text list "Banner_WarnMsg2": 0 '**Local Message Display**'; 1 '~Safety Task Unlocked WB2[0].1'; 2 '~Safety Signature Mismatch WB2[0].2'; 3 '~PLC Battery Bad Or Missing WB2[0].3'; 4 '~Lube System Faulted WB2[0].4'; 5 '~Lube System Cycling WB2[0].5'; 6 '~Lube Level Low WB2[0].6'; 7 '~Spare WB2[0].7'; 8 '~Spare WB2[0].8'; 9 '~Spare WB2[0].9'; 10 '~Main Air Filter Dirty WB2[0].10'; 11 '~Main Water Filter Not OK WB2[0].11'; 12 '~Spare WB2[0].12'; 13 '~Spare WB2[0].13'; 14 '~Spare WB2[0].14'; 15 '~Spare WB2[0].15'; 16 '~Spare WB2[0].16'; 17 '~Spare WB2[0].17'; 18 '~Spare WB2[0].18'; 19 '~Spare WB2[0].19'; 20 '~Spare WB2[0].20'; 21 '~Spare WB2[0].21'; 22 '~Spare WB2[0].22'; 23 '~Spare WB2[0].23'; 24 '~Spare WB2[0].24'; 25 '~Spare WB2[0].25'; 26 '~Spare WB2[0].26'; 27 '~Spare WB2[0].27'; 28 '~Spare WB2[0].28'; 29 '~Spare WB2[0].29'; 30 '~Spare WB2[0].30'; 31 '~Spare WB2[0].31'; 32 '~Sxxx-xxx - Prev Station Exit Lt Scrn Fault - See Prev Station PV WB2[1].0'; 33 '~Sxxx-xxx - Next Station Exit Lt Scrn Fault - See Next Station PV WB2[1].1'; 34 '~Sxxx-xxx - Prev Station Robot In Teach - See Prev Station PV WB2[1].2'; 35 '~Sxxx-xxx - Next Station Robot In Teach - See Next Station PV WB2[1].3'; 36 '~Spare WB2[1].4'; 37 '~Spare WB2[1].5'; 38 '~Sxxx-xxx - Facilities Gate Logic Not Rst - See Facilities Ctrl Pnl WB2[1].6'; 39 '~Spare WB2[1].7'; 40 '~Spare WB2[1].8'; 41 '~Sxxx-xxx - Other Control Zone Fault Present WB2[1].9'; 42 '~Spare WB2[1].10'; 43 '~Spare WB2[1].11'; 44 '~Safety Instruction Warning - Go To Safety Instruction Screen WB2[1].12'; 45 '~Safety Instruction Fault Active - Go To Safety Instuction Screen WB2[1].13'; 46 '~Spare WB2[1].14'; 47 '~Spare WB2[1].15'; 48 '~Spare WB2[1].16'; 49 '~Spare WB2[1].17'; 50 '~Spare WB2[1].18'; 51 '~Spare WB2[1].19'; 52 '~Spare WB2[1].20'; 53 '~Sxxx-xxx Consumed Safety I/O Intlks Not Running-See Source PLC WB2[1].21'; 54 '~Sxxx-xxx Consumed Standard I/O Intlks Not Running-See Source PLC WB2[1].22'; 55 '~Sxxx-xxx Consumed Safety I/O Intlks Not Running-See Source PLC WB2[1].23'; 56 '~Sxxx-xxx Consumed Standard I/O Intlks Not Running-See Source PLC WB2[1].24'; 57 '~Sxxx-xxx Consumed Safety I/O Intlks Not Running-See Source PLC WB2[1].25'; 58 '~Sxxx-xxx Consumed Standard I/O Intlks Not Running-See Source PLC WB2[1].26'; 59 '~Sxxx-xxx Consumed Safety I/O Intlks Not Running-See Source PLC WB2[1].27'; 60 '~Sxxx-xxx Consumed Standard I/O Intlks Not Running-See Source PLC WB2[1].28'; 61 '~Spare WB2[1].29'; 62 '~Spare WB2[1].30'; 63 '~Spare WB2[1].31'; 64 '~Sxxx - xxx E-Stop Depressed - See Station Panel WB2[2].0'; 65 '~Sxxx - xxx E-Stop Circuit Not Reset - Depress Enable Outputs PB WB2[2].1'; 66 '~Sxxx - xxx Safety Gate Open - See Station Panel WB2[2].2'; 67 '~Sxxx - xxx Safety Gate Circuit Not Reset - Depress Gate Reset PB WB2[2].3'; 68 '~Sxxx - xxx Access Or Entry/Exit Light Screen Fault - See Stn Panel WB2[2].4'; 69 '~Sxxx - xxx Robot In Teach - See Station Panel WB2[2].5'; 70 '~Sxxx - xxx Not Ready For Auto - See Station Panel WB2[2].6'; 71 '~Sxxx - xxx Auto Repeat Not Selected - See Station Panel WB2[2].7'; 72 '~Sxxx - xxx Faulted - See Station Panel WB2[2].8'; 73 '~Spare WB2[2].9'; 74 '~Spare WB2[2].10'; 75 '~Spare WB2[2].11'; 76 '~Spare WB2[2].12'; 77 '~Spare WB2[2].13'; 78 '~Spare WB2[2].14'; 79 '~Spare WB2[2].15'; 80 '~Sxxx - xxx E-Stop Depressed - See Station Panel WB2[2].16'; 81 '~Sxxx - xxx E-Stop Circuit Not Reset - Depress Enable Outputs PB WB2[2].17'; 82 '~Sxxx - xxx Safety Gate Open - See Station Panel WB2[2].18'; 83 '~Sxxx - xxx Safety Gate Circuit Not Reset - Depress Gate Reset PB WB2[2].19'; 84 '~Sxxx - xxx Access Or Entry/Exit Light Screen Fault - See Stn Panel WB2[2].20'; 85 '~Sxxx - xxx Robot In Teach - See Station Panel WB2[2].21'; 86 '~Sxxx - xxx Not Ready For Auto - See Station Panel WB2[2].22'; 87 '~Sxxx - xxx Auto Repeat Not Selected - See Station Panel WB2[2].23'; 88 '~Sxxx - xxx Faulted - See Station Panel WB2[2].24'; 89 '~Spare WB2[2].25'; 90 '~Spare WB2[2].26'; 91 '~Spare WB2[2].27'; 92 '~Spare WB2[2].28'; 93 '~Spare WB2[2].29'; 94 '~Spare WB2[2].30'; 95 '~Spare WB2[2].31'; 96 '~Sxxx - xxx E-Stop Depressed - See Station Panel WB2[3].0'; 97 '~Sxxx - xxx E-Stop Circuit Not Reset - Depress Enable Outputs PB WB2[3].1'; 98 '~Sxxx - xxx Safety Gate Open - See Station Panel WB2[3].2'; 99 '~Sxxx - xxx Safety Gate Circuit Not Reset - Depress Gate Reset PB WB2[3].3'; 100 '~Sxxx - xxx Access Or Entry/Exit Light Screen Fault - See Stn Panel WB2[3].4'; 101 '~Sxxx - xxx Robot In Teach - See Station Panel WB2[3].5'; 102 '~Sxxx - xxx Not Ready For Auto - See Station Panel WB2[3].6'; 103 '~Sxxx - xxx Auto Repeat Not Selected - See Station Panel WB2[3].7'; 104 '~Sxxx - xxx Faulted - See Station Panel WB2[3].8'; 105 '~Spare WB2[3].9'; 106 '~Spare WB2[3].10'; 107 '~Spare WB2[3].11'; 108 '~Spare WB2[3].12'; 109 '~Spare WB2[3].13'; 110 '~Spare WB2[3].14'; 111 '~Spare WB2[3].15'; 112 '~Sxxx - xxx E-Stop Depressed - See Station Panel WB2[3].16'; 113 '~Sxxx - xxx E-Stop Circuit Not Reset - Depress Enable Outputs PB WB2[3].17'; 114 '~Sxxx - xxx Safety Gate Open - See Station Panel WB2[3].18'; 115 '~Sxxx - xxx Safety Gate Circuit Not Reset - Depress Gate Reset PB WB2[3].19'; 116 '~Sxxx - xxx Access Or Entry/Exit Light Screen Fault - See Stn Panel WB2[3].20'; 117 '~Sxxx - xxx Robot In Teach - See Station Panel WB2[3].21'; 118 '~Sxxx - xxx Not Ready For Auto - See Station Panel WB2[3].22'; 119 '~Sxxx - xxx Auto Repeat Not Selected - See Station Panel WB2[3].23'; 120 '~Sxxx - xxx Faulted - See Station Panel WB2[3].24'; 121 '~Spare WB2[3].25'; 122 '~Spare WB2[3].26'; 123 '~Spare WB2[3].27'; 124 '~Spare WB2[3].28'; 125 '~Spare WB2[3].29'; 126 '~Spare WB2[3].30'; 127 '~Spare WB2[3].31'; 128 '~Sxxx - xxx E-Stop Depressed - See Station Panel WB2[4].0'; 129 '~Sxxx - xxx E-Stop Circuit Not Reset - Depress Enable Outputs PB WB2[4].1'; 130 '~Sxxx - xxx Safety Gate Open - See Station Panel WB2[4].2'; 131 '~Sxxx - xxx Safety Gate Circuit Not Reset - Depress Gate Reset PB WB2[4].3'; 132 '~Sxxx - xxx Access Or Entry/Exit Light Screen Fault WB2[4].4'; 133 '~Sxxx - xxx Robot In Teach - See Station Panel WB2[4].5'; 134 '~Sxxx - xxx Not Ready For Auto - See Station Panel WB2[4].6'; 135 '~Sxxx - xxx Auto Repeat Not Selected - See Station Panel WB2[4].7'; 136 '~Sxxx - xxx Faulted - See Station Panel WB2[4].8'; 137 '~Spare WB2[4].9'; 138 '~Spare WB2[4].10'; 139 '~Spare WB2[4].11'; 140 '~Spare WB2[4].12'; 141 '~Spare WB2[4].13'; 142 '~Spare WB2[4].14'; 143 '~Spare WB2[4].15'; 144 '~Spare WB2[4].16'; 145 '~Spare WB2[4].17'; 146 '~Spare WB2[4].18'; 147 '~Spare WB2[4].19'; 148 '~Spare WB2[4].20'; 149 '~Spare WB2[4].21'; 150 '~Spare WB2[4].22'; 151 '~Spare WB2[4].23'; 152 '~Spare WB2[4].24'; 153 '~Spare WB2[4].25'; 154 '~Spare WB2[4].26'; 155 '~Spare WB2[4].27'; 156 '~Spare WB2[4].28'; 157 '~Spare WB2[4].29'; 158 '~Spare WB2[4].30'; 159 '~Spare WB2[4].31'; 160 '~S002 Safety Gate Logic Not Reset - Depress Gate Reset PB WB2[5].0'; 161 '~Spare WB2[5].1'; 162 '~Spare WB2[5].2'; 163 '~Spare WB2[5].3'; 164 '~S002 Ready For Automatic Depress Auto PB WB2[5].4'; 165 '~S002 Master Logic Not Reset Depress Enable Ouputs PB WB2[5].5'; 166 '~S002 Not Ready For Automatic WB2[5].6'; 167 '~S002 Auto Repeat Not Selected - See Utility Screen WB2[5].7'; 168 '~Spare WB2[5].8'; 169 '~Spare WB2[5].9'; 170 '~S002 Service Side Light Screen Not Reset - Depress Cycle Start PB WB2[5].10'; 171 '~S002 Remote Side Light Screen Not Reset - Depress Cycle Start PB WB2[5].11'; 172 '~Spare WB2[5].12'; 173 '~Spare WB2[5].13'; 174 '~Spare WB2[5].14'; 175 '~Spare WB2[5].15'; 176 '~Spare WB2[5].16'; 177 '~Spare WB2[5].17'; 178 '~Spare WB2[5].18'; 179 '~Spare WB2[5].19'; 180 '~Spare WB2[5].20'; 181 '~Spare WB2[5].21'; 182 '~Spare WB2[5].22'; 183 '~Spare WB2[5].23'; 184 '~S002 Service Side Model 1 Prycheck Selected WB2[5].24'; 185 '~S002 Remote Side Model 1 Prycheck Selected WB2[5].25'; 186 '~S002 Service Side Model 2 Prycheck Selected WB2[5].26'; 187 '~S002 Remote Side Model 2 Prycheck Selected WB2[5].27'; 188 '~Spare WB2[5].28'; 189 '~Spare WB2[5].29'; 190 '~Spare WB2[5].30'; 191 '~Spare WB2[5].31'; 192 '~Spare WB2[6].0'; 193 '~Spare WB2[6].1'; 194 '~S002 Oper #1 Light Screen Not Reset - Press Cycle Start PB WB2[6].2'; 195 '~S002 Oper #2 Light Screen Not Reset - Press Cycle Start PB WB2[6].3'; 196 '~S002CV# Oper #1 Lt Screen Not Reset - Press Cycle Start PB WB2[6].4'; 197 '~S002CV# Oper #2 Lt Screen Not Reset - Press Cycle Start PB WB2[6].5'; 198 '~Spare WB2[6].6'; 199 '~Spare WB2[6].7'; 200 '~Spare WB2[6].8'; 201 '~Spare WB2[6].9'; 202 '~S002 Operator #1 Cycle Over Time WB2[6].10'; 203 '~S002 Operator #2 Cycle Overtime WB2[6].11'; 204 '~S002TT1 Operator #1 Cycle Over Time WB2[6].12'; 205 '~S003TL1 Operator #1 Cycle Over Time WB2[6].13'; 206 '~Spare WB2[6].14'; 207 '~Spare WB2[6].15'; 208 '~Spare WB2[6].16'; 209 '~Spare WB2[6].17'; 210 '~Spare WB2[6].18'; 211 '~Spare WB2[6].19'; 212 '~Spare WB2[6].20'; 213 '~Spare WB2[6].21'; 214 '~Spare WB2[6].22'; 215 '~Spare WB2[6].23'; 216 '~Spare WB2[6].24'; 217 '~Spare WB2[6].25'; 218 '~Spare WB2[6].26'; 219 '~Spare WB2[6].27'; 220 '~Spare WB2[6].28'; 221 '~Spare WB2[6].29'; 222 '~Spare WB2[6].30'; 223 '~Spare WB2[6].31'; 224 '~PDPES1 - PDP EtherNet Switch Port At Half Duplex WB2[7].0'; 225 '~PDPES1 - PDP EtherNet Switch Configuration Changes Not Saved WB2[7].1'; 226 '~PDPES1 - PDP EtherNet Switch Configuration Changed WB2[7].2'; 227 '~PDPES1 - PDP EtherNet Switch Port With Excessive Errors WB2[7].3'; 228 '~PDPES1 - PDP EtherNet Switch Port With Utilization Warning WB2[7].4'; 229 '~PDPES1 - PDP EtherNet Switch Changes Require Reboot WB2[7].5'; 230 '~Spare WB2[7].6'; 231 '~Spare WB2[7].7'; 232 '~MPES1 - Main Panel EtherNet Switch Port At Half Duplex WB2[7].8'; 233 '~MPES1 - Main Panel EtherNet Switch Configuration Changes Not Saved WB2[7].9'; 234 '~MPES1 - Main Panel EtherNet Switch Configuration Changed WB2[7].10'; 235 '~MPES1 - Main Panel EtherNet Switch Port With Excessive Errors WB2[7].11'; 236 '~MPES1 - Main Panel EtherNet Switch Port With Utilization Warning WB2[7].12'; 237 '~MPES1 - Main Panel EtherNet Switch Changes Require Reboot WB2[7].13'; 238 '~Spare WB2[7].14'; 239 '~Spare WB2[7].15'; 240 '~MPES2 - Main Panel EtherNet Switch Port At Half Duplex WB2[7].16'; 241 '~MPES2 - Main Panel EtherNet Switch Configuration Changes Not Saved WB2[7].17'; 242 '~MPES2 - Main Panel EtherNet Switch Configuration Changed WB2[7].18'; 243 '~MPES2 - Main Panel EtherNet Switch Port With Excessive Errors WB2[7].19'; 244 '~MPES2 - Main Panel EtherNet Switch Port With Utilization Warning WB2[7].20'; 245 '~MPES2 - Main Panel EtherNet Switch Changes Require Reboot WB2[7].21'; 246 '~Spare WB2[7].22'; 247 '~Spare WB2[7].23'; 248 '~MPES3 - Main Panel EtherNet Switch Port At Half Duplex WB2[7].24'; 249 '~MPES3 - Main Panel EtherNet Switch Configuration Changes Not Saved WB2[7].25'; 250 '~MPES3 - Main Panel EtherNet Switch Configuration Changed WB2[7].26'; 251 '~MPES3 - Main Panel EtherNet Switch Port With Excessive Errors WB2[7].27'; 252 '~MPES3 - Main Panel EtherNet Switch Port With Utilization Warning WB2[7].28'; 253 '~MPES3 - Main Panel EtherNet Switch Changes Require Reboot WB2[7].29'; 254 '~Spare WB2[7].30'; 255 '~Spare WB2[7].31'; 256 '~PV3ES1 - PV3 EtherNet Switch Port At Half Duplex WB2[8].0'; 257 '~PV3ES1 - PV3 EtherNet Switch Configuration Changes Not Saved WB2[8].1'; 258 '~PV3ES1 - PV3 EtherNet Switch Configuration Changed WB2[8].2'; 259 '~PV3ES1 - PV3 EtherNet Switch Port With Excessive Errors WB2[8].3'; 260 '~PV3ES1 - PV3 EtherNet Switch Port With Utilization Warning WB2[8].4'; 261 '~PV3ES1 - PV3 EtherNet Switch Changes Require Reboot WB2[8].5'; 262 '~Spare WB2[8].6'; 263 '~Spare WB2[8].7'; 264 '~PV4ES1 - PV4 EtherNet Switch Port At Half Duplex WB2[8].8'; 265 '~PV4ES1 - PV4 EtherNet Switch Configuration Changes Not Saved WB2[8].9'; 266 '~PV4ES1 - PV4 EtherNet Switch Configuration Changed WB2[8].10'; 267 '~PV4ES1 - PV4 EtherNet Switch Port With Excessive Errors WB2[8].11'; 268 '~PV4ES1 - PV4 EtherNet Switch Port With Utilization Warning WB2[8].12'; 269 '~PV4ES1 - PV4 EtherNet Switch Changes Require Reboot WB2[8].13'; 270 '~Spare WB2[8].14'; 271 '~Spare WB2[8].15'; 272 '~ES3ES1 - ES3 EtherNet Switch Port At Half Duplex WB2[8].16'; 273 '~ES3ES1 - ES3 EtherNet Switch Configuration Changes Not Saved WB2[8].17'; 274 '~ES3ES1 - ES3 EtherNet Switch Configuration Changed WB2[8].18'; 275 '~ES3ES1 - ES3 EtherNet Switch Port With Excessive Errors WB2[8].19'; 276 '~ES3ES1 - ES3 EtherNet Switch Port With Utilization Warning WB2[8].20'; 277 '~ES3ES1 - ES3 EtherNet Switch Changes Require Reboot WB2[8].21'; 278 '~Spare WB2[8].22'; 279 '~Spare WB2[8].23'; 280 '~ES4ES1 - ES4 EtherNet Switch Port At Half Duplex WB2[8].24'; 281 '~ES4ES1 - ES4 EtherNet Switch Configuration Changes Not Saved WB2[8].25'; 282 '~ES4ES1 - ES4 EtherNet Switch Configuration Changed WB2[8].26'; 283 '~ES4ES1 - ES4 EtherNet Switch Port With Excessive Errors WB2[8].27'; 284 '~ES4ES1 - ES4 EtherNet Switch Port With Utilization Warning WB2[8].28'; 285 '~ES4ES1 - ES4 EtherNet Switch Changes Require Reboot WB2[8].29'; 286 '~Spare WB2[8].30'; 287 '~Spare WB2[8].31'; 288 '~Spare WB2[9].0'; 289 '~Spare WB2[9].1'; 290 '~Spare WB2[9].2'; 291 '~Spare WB2[9].3'; 292 '~Spare WB2[9].4'; 293 '~Spare WB2[9].5'; 294 '~Spare WB2[9].6'; 295 '~Spare WB2[9].7'; 296 '~Spare WB2[9].8'; 297 '~Spare WB2[9].9'; 298 '~Spare WB2[9].10'; 299 '~Spare WB2[9].11'; 300 '~Spare WB2[9].12'; 301 '~Spare WB2[9].13'; 302 '~Spare WB2[9].14'; 303 '~Spare WB2[9].15'; 304 '~Spare WB2[9].16'; 305 '~Spare WB2[9].17'; 306 '~Spare WB2[9].18'; 307 '~Spare WB2[9].19'; 308 '~Spare WB2[9].20'; 309 '~Spare WB2[9].21'; 310 '~Spare WB2[9].22'; 311 '~Spare WB2[9].23'; 312 '~Spare WB2[9].24'; 313 '~Spare WB2[9].25'; 314 '~Spare WB2[9].26'; 315 '~Spare WB2[9].27'; 316 '~Spare WB2[9].28'; 317 '~Spare WB2[9].29'; 318 '~Spare WB2[9].30'; 319 '~Spare WB2[9].31'; 320 '~S001R09 Waiting Zone #1 Not Clear WB2[10].0'; 321 '~S001R09 Waiting Zone #2 Not Clear WB2[10].1'; 322 '~S001R09 Waiting Zone #3 Not Clear WB2[10].2'; 323 '~S001R09 Waiting Zone #4 Not Clear WB2[10].3'; 324 '~S001R09 Waiting Zone #5 Not Clear WB2[10].4'; 325 '~S001R09 Waiting Zone #6 Not Clear WB2[10].5'; 326 '~S001R09 Waiting Zone #7 Not Clear WB2[10].6'; 327 '~S001R09 Waiting Zone #8 Not Clear WB2[10].7'; 328 '~S001R09 Waiting Zone #9 Not Clear WB2[10].8'; 329 '~S001R09 Waiting Zone #10 Not Clear WB2[10].9'; 330 '~S001R09 Waiting Zone #11 Not Clear WB2[10].10'; 331 '~S001R09 Waiting Zone #12 Not Clear WB2[10].11'; 332 '~S001R09 Waiting Zone #13 Not Clear WB2[10].12'; 333 '~S001R09 Waiting Zone #14 Not Clear WB2[10].13'; 334 '~S001R09 Waiting Tip Dress Zone #1 Not Clear WB2[10].14'; 335 '~S001R09 Waiting Tip Dress Zone #2 Not Clear WB2[10].15'; 336 '~S001R09 Adjacent Robot xx-xx In Teach WB2[10].16'; 337 '~S001R09 Adjacent Robot xx-xx In Teach WB2[10].17'; 338 '~S001R09 Adjacent Robot xx-xx In Teach WB2[10].18'; 339 '~S001R09 Adjacent Robot xx-xx In Teach WB2[10].19'; 340 '~S001R09 Adjacent Robot xx-xx In Teach WB2[10].20'; 341 '~S001R09 Adjacent Robot xx-xx In Teach WB2[10].21'; 342 '~S001R09 Adjacent Robot xx-xx In Teach WB2[10].22'; 343 '~S001R09 Adjacent Robot xx-xx In Teach WB2[10].23'; 344 '~S001R09 Adjacent Robot xx-xx In Teach WB2[10].24'; 345 '~S001R09 Adjacent Robot xx-xx In Teach WB2[10].25'; 346 '~Spare WB2[10].26'; 347 '~Spare WB2[10].27'; 348 '~Spare WB2[10].28'; 349 '~S001R09 Robot Not Clear Of Fixture WB2[10].29'; 350 '~Spare WB2[10].30'; 351 '~Spare WB2[10].31'; 352 '~Spare WB2[11].0'; 353 '~Spare WB2[11].1'; 354 '~Spare WB2[11].2'; 355 '~Spare WB2[11].3'; 356 '~Spare WB2[11].4'; 357 '~Spare WB2[11].5'; 358 '~Spare WB2[11].6'; 359 '~Spare WB2[11].7'; 360 '~Spare WB2[11].8'; 361 '~Spare WB2[11].9'; 362 '~Spare WB2[11].10'; 363 '~Spare WB2[11].11'; 364 '~Spare WB2[11].12'; 365 '~Spare WB2[11].13'; 366 '~Spare WB2[11].14'; 367 '~Spare WB2[11].15'; 368 '~Spare WB2[11].16'; 369 '~Spare WB2[11].17'; 370 '~Spare WB2[11].18'; 371 '~Spare WB2[11].19'; 372 '~Spare WB2[11].20'; 373 '~Spare WB2[11].21'; 374 '~Spare WB2[11].22'; 375 '~Spare WB2[11].23'; 376 '~Spare WB2[11].24'; 377 '~Spare WB2[11].25'; 378 '~Spare WB2[11].26'; 379 '~Spare WB2[11].27'; 380 '~Spare WB2[11].28'; 381 '~Spare WB2[11].29'; 382 '~Spare WB2[11].30'; 383 '~Spare WB2[11].31'; 384 '~S001R09 Cycle Overtime WB2[12].0'; 385 '~S001R09 In Bypass WB2[12].1'; 386 '~S001R09 Battery Low WB2[12].2'; 387 '~S001R09 Servo Over Torque WB2[12].3'; 388 '~S001R09 Process Retry In Progress WB2[12].4'; 389 '~Spare WB2[12].5'; 390 '~S001R09 Robot Edit Occurred Ext App WB2[12].6'; 391 '~S001R09 Robot Input Simmed WB2[12].7'; 392 '~S001R09 Robot Output Simmed WB2[12].8'; 393 '~Spare WB2[12].9'; 394 '~Spare WB2[12].10'; 395 '~Spare WB2[12].11'; 396 '~Spare WB2[12].12'; 397 '~Spare WB2[12].13'; 398 '~Spare WB2[12].14'; 399 '~Spare WB2[12].15'; 400 '~S001R09F1B1.M.ModuleFlt - Externa App 1 I/O Module Warning WB2[12].16'; 401 '~S001R09F2B1.M.ModuleFlt - Externa App 2 I/O Module Warning WB2[12].17'; 402 '~S001R09F3B1.M.ModuleFlt - Externa App 3 I/O Module Warning WB2[12].18'; 403 '~Spare WB2[12].19'; 404 '~Spare WB2[12].20'; 405 '~Spare WB2[12].21'; 406 '~Spare WB2[12].22'; 407 '~Spare WB2[12].23'; 408 '~S001R09ES1 - S001R09 EtherNet Switch Port At Half Duplex WB2[12].24'; 409 '~S001R09ES1 - S001R09 EtherNet Switch Config Changes Not Saved WB2[12].25'; 410 '~S001R09ES1 - S001R09 EtherNet Switch Configuration Changed WB2[12].26'; 411 '~S001R09ES1 - S001R09 EtherNet Switch Port With Excessive Errors WB2[12].27'; 412 '~S001R09ES1 - S001R09 EtherNet Switch Port With Utilization Warning WB2[12].28'; 413 '~S001R09ES1 - S001R09 EtherNet Switch Changes Require Reboot WB2[12].29'; 414 '~Spare WB2[12].30'; 415 '~Spare WB2[12].31'; 416 '~Spare WB2[13].0'; 417 '~Spare WB2[13].1'; 418 '~S001R09 Servo Gun Tip Calib Request 1 WB2[13].2'; 419 '~S001R09 I-Available Warning 1 WB2[13].3'; 420 '~S001R09 Tip Dress Motor 1 Fault Bypassed WB2[13].4'; 421 '~S001R09 Tip Change Notice 1 WB2[13].5'; 422 '~S001R09 Bypass Tip Dresser 1 Selected WB2[13].6'; 423 '~S001R09 Auto Tip Changer Low 1 WB2[13].7'; 424 '~S001R09 Auto Tip Changer Empty 1 WB2[13].8'; 425 '~S001R09 Tip Wear Ratio Warning 1 - Touch Up Tip Dress Program WB2[13].9'; 426 '~S001R09 Stud Weld 1 Maintenance Reqd WB2[13].10'; 427 '~S001R09 Stud Weld 1 Low Stud Warning WB2[13].11'; 428 '~Spare WB2[13].12'; 429 '~S001R09 Rivet 1 Low Rivet Warning WB2[13].13'; 430 '~S001R09 Rivet 1 - Skip Once Initiated from Robot TP WB2[13].14'; 431 '~S001R09 Rivet 1 - Skip Remaining Initiated from Robot TP WB2[13].15'; 432 '~S001R09 Rivet 1 Preventive Maintenace Required WB2[13].16'; 433 '~S001R09 Rivet 1 Magazine Low WB2[13].17'; 434 '~S001R09 Tip Change 1 Bypassed WB2[13].18'; 435 '~S001R09 Mig Weld Fluid Level Low WB2[13].19'; 436 '~S001R09 Weld Ctrlr 1 Adaptive Mode Is Disabled WB2[13].20'; 437 '~S001R09 Tip Cutter 1 Warning WB2[13].21'; 438 '~S001R09 Rivet 1 Tape-Cut Required WB2[13].22'; 439 '~S001R09 Wire Feeder Motor Over Current WB2[13].23'; 440 '~Spare WB2[13].24'; 441 '~S001R09 Sealer Ctrlr 1 Minor Fault WB2[13].25'; 442 '~S001R09 Sealer Ctrlr 1 Required Rezeroing WB2[13].26'; 443 '~S001R09 Loaded To Average WB2[13].27'; 444 '~S001R09 Vision Process Aborted WB2[13].28'; 445 '~S001R09 Vision System Trending WB2[13].29'; 446 '~S001R09 Vision Out Of Tolerance WB2[13].30'; 447 '~Spare WB2[13].31'; 448 '~Spare WB2[14].0'; 449 '~Spare WB2[14].1'; 450 '~S001R09 Servo Gun Tip Calib Request 2 WB2[14].2'; 451 '~S001R09 I-Available Warning 2 WB2[14].3'; 452 '~S001R09 Tip Dress Motor 2 Fault Bypassed WB2[14].4'; 453 '~S001R09 Tip Change Notice 2 WB2[14].5'; 454 '~S001R09 Bypass Tip Dresser 2 Selected WB2[14].6'; 455 '~S001R09 Auto Tip Changer Low 2 WB2[14].7'; 456 '~S001R09 Auto Tip Changer Empty 2 WB2[14].8'; 457 '~S001R09 Tip Wear Ratio Warning 2 - Touch Up Tip Dress Program WB2[14].9'; 458 '~S001R09 Stud Weld 2 Maintenance Reqd WB2[14].10'; 459 '~S001R09 Stud Weld 2 Low Stud Warning WB2[14].11'; 460 '~Spare WB2[14].12'; 461 '~S001R09 Rivet 2 Low Rivet Warning WB2[14].13'; 462 '~S001R09 Rivet 2 - Skip Once Initiated from Robot TP WB2[14].14'; 463 '~S001R09 Rivet 2 - Skip Remaining Initiated from Robot TP WB2[14].15'; 464 '~S001R09 Rivet 2 Preventive Maintenace Required WB2[14].16'; 465 '~S001R09 Rivet 2 Magazine Low WB2[14].17'; 466 '~S001R09 Tip Change 2 Bypassed WB2[14].18'; 467 '~S001R09 Laser Dirty Glass Warning WB2[14].19'; 468 '~S001R09 Weld Ctrlr 2 Adaptive Mode Is Disabled WB2[14].20'; 469 '~S001R09 Tip Cutter 2 Warning WB2[14].21'; 470 '~S001R09 Rivet 2 Tape-Cut Required WB2[14].22'; 471 '~S001R09 Mig Tip Nozzel Replacement Warning WB2[14].23'; 472 '~S001R09 Mig Tip Nozzel Replacement Required WB2[14].24'; 473 '~S001R09 Sealer Ctrlr 2 Minor Fault WB2[14].25'; 474 '~S001R09 Sealer Ctrlr 2 Required Rezeroing WB2[14].26'; 475 '~S001R09 Mig Barrel Replacement Warning WB2[14].27'; 476 '~S001R09 Mig Barrel Replacement Required WB2[14].28'; 477 '~S001R09 In Touch Up Mode WB2[14].29'; 478 '~S001R09 Touch Up Mode Not Enabled WB2[14].30'; 479 '~Spare WB2[14].31'; 480 '~S001R09 Laser Controller Fault WB2[15].0'; 481 '~S001R09 Laser Dirty Glass Warning WB2[15].1'; 482 '~S001R09 Laser Warning WB2[15].2'; 483 '~Spare WB2[15].3'; 484 '~Spare WB2[15].4'; 485 '~Spare WB2[15].5'; 486 '~Spare WB2[15].6'; 487 '~Spare WB2[15].7'; 488 '~Spare WB2[15].8'; 489 '~Spare WB2[15].9'; 490 '~Spare WB2[15].10'; 491 '~Spare WB2[15].11'; 492 '~Spare WB2[15].12'; 493 '~Spare WB2[15].13'; 494 '~Spare WB2[15].14'; 495 '~Spare WB2[15].15'; 496 '~Spare WB2[15].16'; 497 '~Spare WB2[15].17'; 498 '~Spare WB2[15].18'; 499 '~Spare WB2[15].19'; 500 '~Spare WB2[15].20'; 501 '~Spare WB2[15].21'; 502 '~Spare WB2[15].22'; 503 '~Spare WB2[15].23'; 504 '~Spare WB2[15].24'; 505 '~Spare WB2[15].25'; 506 '~Spare WB2[15].26'; 507 '~Spare WB2[15].27'; 508 '~Spare WB2[15].28'; 509 '~Spare WB2[15].29'; 510 '~Spare WB2[15].30'; 511 '~Spare WB2[15].31'; 512 '~Spare WB2[16].0'; 513 '~Spare WB2[16].1'; 514 '~Spare WB2[16].2'; 515 '~Spare WB2[16].3'; 516 '~Spare WB2[16].4'; 517 '~Spare WB2[16].5'; 518 '~Spare WB2[16].6'; 519 '~Spare WB2[16].7'; 520 '~Spare WB2[16].8'; 521 '~Spare WB2[16].9'; 522 '~Spare WB2[16].10'; 523 '~Spare WB2[16].11'; 524 '~Spare WB2[16].12'; 525 '~Spare WB2[16].13'; 526 '~Spare WB2[16].14'; 527 '~Spare WB2[16].15'; 528 '~Spare WB2[16].16'; 529 '~Spare WB2[16].17'; 530 '~Spare WB2[16].18'; 531 '~Spare WB2[16].19'; 532 '~Spare WB2[16].20'; 533 '~Spare WB2[16].21'; 534 '~Spare WB2[16].22'; 535 '~Spare WB2[16].23'; 536 '~Spare WB2[16].24'; 537 '~Spare WB2[16].25'; 538 '~Spare WB2[16].26'; 539 '~Spare WB2[16].27'; 540 '~Spare WB2[16].28'; 541 '~Spare WB2[16].29'; 542 '~Spare WB2[16].30'; 543 '~Spare WB2[16].31'; 544 '~Spare WB2[17].0'; 545 '~Spare WB2[17].1'; 546 '~Spare WB2[17].2'; 547 '~Spare WB2[17].3'; 548 '~Spare WB2[17].4'; 549 '~Spare WB2[17].5'; 550 '~Spare WB2[17].6'; 551 '~Spare WB2[17].7'; 552 '~Spare WB2[17].8'; 553 '~Spare WB2[17].9'; 554 '~Spare WB2[17].10'; 555 '~Spare WB2[17].11'; 556 '~Spare WB2[17].12'; 557 '~Spare WB2[17].13'; 558 '~Spare WB2[17].14'; 559 '~Spare WB2[17].15'; 560 '~Spare WB2[17].16'; 561 '~Spare WB2[17].17'; 562 '~Spare WB2[17].18'; 563 '~Spare WB2[17].19'; 564 '~Spare WB2[17].20'; 565 '~Spare WB2[17].21'; 566 '~Spare WB2[17].22'; 567 '~Spare WB2[17].23'; 568 '~Spare WB2[17].24'; 569 '~Spare WB2[17].25'; 570 '~Spare WB2[17].26'; 571 '~Spare WB2[17].27'; 572 '~Spare WB2[17].28'; 573 '~Spare WB2[17].29'; 574 '~Spare WB2[17].30'; 575 '~Spare WB2[17].31'; 576 '~S001R10 Waiting Zone #1 Not Clear WB2[18].0'; 577 '~S001R10 Waiting Zone #2 Not Clear WB2[18].1'; 578 '~S001R10 Waiting Zone #3 Not Clear WB2[18].2'; 579 '~S001R10 Waiting Zone #4 Not Clear WB2[18].3'; 580 '~S001R10 Waiting Zone #5 Not Clear WB2[18].4'; 581 '~S001R10 Waiting Zone #6 Not Clear WB2[18].5'; 582 '~S001R10 Waiting Zone #7 Not Clear WB2[18].6'; 583 '~S001R10 Waiting Zone #8 Not Clear WB2[18].7'; 584 '~S001R10 Waiting Zone #9 Not Clear WB2[18].8'; 585 '~S001R10 Waiting Zone #10 Not Clear WB2[18].9'; 586 '~S001R10 Waiting Zone #11 Not Clear WB2[18].10'; 587 '~S001R10 Waiting Zone #12 Not Clear WB2[18].11'; 588 '~S001R10 Waiting Zone #13 Not Clear WB2[18].12'; 589 '~S001R10 Waiting Zone #14 Not Clear WB2[18].13'; 590 '~S001R10 Waiting Tip Dress Zone #1 Not Clear WB2[18].14'; 591 '~S001R10 Waiting Tip Dress Zone #2 Not Clear WB2[18].15'; 592 '~S001R10 Adjacent Robot xx-xx In Teach WB2[18].16'; 593 '~S001R10 Adjacent Robot xx-xx In Teach WB2[18].17'; 594 '~S001R10 Adjacent Robot xx-xx In Teach WB2[18].18'; 595 '~S001R10 Adjacent Robot xx-xx In Teach WB2[18].19'; 596 '~S001R10 Adjacent Robot xx-xx In Teach WB2[18].20'; 597 '~S001R10 Adjacent Robot xx-xx In Teach WB2[18].21'; 598 '~S001R10 Adjacent Robot xx-xx In Teach WB2[18].22'; 599 '~S001R10 Adjacent Robot xx-xx In Teach WB2[18].23'; 600 '~S001R10 Adjacent Robot xx-xx In Teach WB2[18].24'; 601 '~S001R10 Adjacent Robot xx-xx In Teach WB2[18].25'; 602 '~Spare WB2[18].26'; 603 '~Spare WB2[18].27'; 604 '~Spare WB2[18].28'; 605 '~S001R10 Robot Not Clear Of Fixture WB2[18].29'; 606 '~Spare WB2[18].30'; 607 '~Spare WB2[18].31'; 608 '~Spare WB2[19].0'; 609 '~Spare WB2[19].1'; 610 '~Spare WB2[19].2'; 611 '~Spare WB2[19].3'; 612 '~Spare WB2[19].4'; 613 '~Spare WB2[19].5'; 614 '~Spare WB2[19].6'; 615 '~Spare WB2[19].7'; 616 '~Spare WB2[19].8'; 617 '~Spare WB2[19].9'; 618 '~Spare WB2[19].10'; 619 '~Spare WB2[19].11'; 620 '~Spare WB2[19].12'; 621 '~Spare WB2[19].13'; 622 '~Spare WB2[19].14'; 623 '~Spare WB2[19].15'; 624 '~Spare WB2[19].16'; 625 '~Spare WB2[19].17'; 626 '~Spare WB2[19].18'; 627 '~Spare WB2[19].19'; 628 '~Spare WB2[19].20'; 629 '~Spare WB2[19].21'; 630 '~Spare WB2[19].22'; 631 '~Spare WB2[19].23'; 632 '~Spare WB2[19].24'; 633 '~Spare WB2[19].25'; 634 '~Spare WB2[19].26'; 635 '~Spare WB2[19].27'; 636 '~Spare WB2[19].28'; 637 '~Spare WB2[19].29'; 638 '~Spare WB2[19].30'; 639 '~Spare WB2[19].31'; 640 '~S001R10 Cycle Overtime WB2[20].0'; 641 '~S001R10 In Bypass WB2[20].1'; 642 '~S001R10 Battery Low WB2[20].2'; 643 '~S001R10 Servo Over Torque WB2[20].3'; 644 '~S001R10 Process Retry In Progress WB2[20].4'; 645 '~Spare WB2[20].5'; 646 '~S001R10 Robot Edit Occurred Ext App WB2[20].6'; 647 '~S001R10 Robot Input Simmed WB2[20].7'; 648 '~S001R10 Robot Output Simmed WB2[20].8'; 649 '~Spare WB2[20].9'; 650 '~Spare WB2[20].10'; 651 '~Spare WB2[20].11'; 652 '~Spare WB2[20].12'; 653 '~Spare WB2[20].13'; 654 '~Spare WB2[20].14'; 655 '~Spare WB2[20].15'; 656 '~S001R10F1B1.M.ModuleFlt - Externa App 1 I/O Module Warning WB2[20].16'; 657 '~S001R10F2B1.M.ModuleFlt - Externa App 2 I/O Module Warning WB2[20].17'; 658 '~S001R10F3B1.M.ModuleFlt - Externa App 3 I/O Module Warning WB2[20].18'; 659 '~Spare WB2[20].19'; 660 '~Spare WB2[20].20'; 661 '~Spare WB2[20].21'; 662 '~Spare WB2[20].22'; 663 '~Spare WB2[20].23'; 664 '~S001R10ES1 - S001R10 EtherNet Switch Port At Half Duplex WB2[20].24'; 665 '~S001R10ES1 - S001R10 EtherNet Switch Config Changes Not Saved WB2[20].25'; 666 '~S001R10ES1 - S001R10 EtherNet Switch Configuration Changed WB2[20].26'; 667 '~S001R10ES1 - S001R10 EtherNet Switch Port With Excessive Errors WB2[20].27'; 668 '~S001R10ES1 - S001R10 EtherNet Switch Port With Utilization Warning WB2[20].28'; 669 '~S001R10ES1 - S001R10 EtherNet Switch Changes Require Reboot WB2[20].29'; 670 '~Spare WB2[20].30'; 671 '~Spare WB2[20].31'; 672 '~Spare WB2[21].0'; 673 '~Spare WB2[21].1'; 674 '~S001R10 Servo Gun Tip Calib Request 1 WB2[21].2'; 675 '~S001R10 I-Available Warning 1 WB2[21].3'; 676 '~S001R10 Tip Dress Motor 1 Fault Bypassed WB2[21].4'; 677 '~S001R10 Tip Change Notice 1 WB2[21].5'; 678 '~S001R10 Bypass Tip Dresser 1 Selected WB2[21].6'; 679 '~S001R10 Auto Tip Changer Low 1 WB2[21].7'; 680 '~S001R10 Auto Tip Changer Empty 1 WB2[21].8'; 681 '~S001R10 Tip Wear Ratio Warning 1 - Touch Up Tip Dress Program WB2[21].9'; 682 '~S001R10 Stud Weld 1 Maintenance Reqd WB2[21].10'; 683 '~S001R10 Stud Weld 1 Low Stud Warning WB2[21].11'; 684 '~Spare WB2[21].12'; 685 '~S001R10 Rivet 1 Low Rivet Warning WB2[21].13'; 686 '~S001R10 Rivet 1 - Skip Once Initiated from Robot TP WB2[21].14'; 687 '~S001R10 Rivet 1 - Skip Remaining Initiated from Robot TP WB2[21].15'; 688 '~S001R10 Rivet 1 Preventive Maintenace Required WB2[21].16'; 689 '~S001R10 Rivet 1 Magazine Low WB2[21].17'; 690 '~S001R10 Tip Change 1 Bypassed WB2[21].18'; 691 '~S001R10 Mig Weld Fluid Level Low WB2[21].19'; 692 '~S001R10 Weld Ctrlr 1 Adaptive Mode Is Disabled WB2[21].20'; 693 '~S001R10 Tip Cutter 1 Warning WB2[21].21'; 694 '~S001R10 Rivet 1 Tape-Cut Required WB2[21].22'; 695 '~S001R10 Wire Feeder Motor Over Current WB2[21].23'; 696 '~Spare WB2[21].24'; 697 '~S001R10 Sealer Ctrlr 1 Minor Fault WB2[21].25'; 698 '~S001R10 Sealer Ctrlr 1 Required Rezeroing WB2[21].26'; 699 '~S001R10 Loaded To Average WB2[21].27'; 700 '~S001R10 Vision Process Aborted WB2[21].28'; 701 '~S001R10 Vision System Trending WB2[21].29'; 702 '~S001R10 Vision Out Of Tolerance WB2[21].30'; 703 '~Spare WB2[21].31'; 704 '~Spare WB2[22].0'; 705 '~Spare WB2[22].1'; 706 '~S001R10 Servo Gun Tip Calib Request 2 WB2[22].2'; 707 '~S001R10 I-Available Warning 2 WB2[22].3'; 708 '~S001R10 Tip Dress Motor 2 Fault Bypassed WB2[22].4'; 709 '~S001R10 Tip Change Notice 2 WB2[22].5'; 710 '~S001R10 Bypass Tip Dresser 2 Selected WB2[22].6'; 711 '~S001R10 Auto Tip Changer Low 2 WB2[22].7'; 712 '~S001R10 Auto Tip Changer Empty 2 WB2[22].8'; 713 '~S001R10 Tip Wear Ratio Warning 2 - Touch Up Tip Dress Program WB2[22].9'; 714 '~S001R10 Stud Weld 2 Maintenance Reqd WB2[22].10'; 715 '~S001R10 Stud Weld 2 Low Stud Warning WB2[22].11'; 716 '~Spare WB2[22].12'; 717 '~S001R10 Rivet 2 Low Rivet Warning WB2[22].13'; 718 '~S001R10 Rivet 2 - Skip Once Initiated from Robot TP WB2[22].14'; 719 '~S001R10 Rivet 2 - Skip Remaining Initiated from Robot TP WB2[22].15'; 720 '~S001R10 Rivet 2 Preventive Maintenace Required WB2[22].16'; 721 '~S001R10 Rivet 2 Magazine Low WB2[22].17'; 722 '~S001R10 Tip Change 2 Bypassed WB2[22].18'; 723 '~S001R10 Laser Dirty Glass Warning WB2[22].19'; 724 '~S001R10 Weld Ctrlr 2 Adaptive Mode Is Disabled WB2[22].20'; 725 '~S001R10 Tip Cutter 2 Warning WB2[22].21'; 726 '~S001R10 Rivet 2 Tape-Cut Required WB2[22].22'; 727 '~S001R10 Mig Tip Nozzel Replacement Warning WB2[22].23'; 728 '~S001R10 Mig Tip Nozzel Replacement Required WB2[22].24'; 729 '~S001R10 Sealer Ctrlr 2 Minor Fault WB2[22].25'; 730 '~S001R10 Sealer Ctrlr 2 Required Rezeroing WB2[22].26'; 731 '~S001R10 Mig Barrel Replacement Warning WB2[22].27'; 732 '~S001R10 Mig Barrel Replacement Required WB2[22].28'; 733 '~S001R10 In Touch Up Mode WB2[22].29'; 734 '~S001R10 Touch Up Mode Not Enabled WB2[22].30'; 735 '~Spare WB2[22].31'; 736 '~S001R10 Laser Controller Fault WB2[23].0'; 737 '~S001R10 Laser Dirty Glass Warning WB2[23].1'; 738 '~S001R10 Laser Warning WB2[23].2'; 739 '~Spare WB2[23].3'; 740 '~Spare WB2[23].4'; 741 '~Spare WB2[23].5'; 742 '~Spare WB2[23].6'; 743 '~Spare WB2[23].7'; 744 '~Spare WB2[23].8'; 745 '~Spare WB2[23].9'; 746 '~Spare WB2[23].10'; 747 '~Spare WB2[23].11'; 748 '~Spare WB2[23].12'; 749 '~Spare WB2[23].13'; 750 '~Spare WB2[23].14'; 751 '~Spare WB2[23].15'; 752 '~Spare WB2[23].16'; 753 '~Spare WB2[23].17'; 754 '~Spare WB2[23].18'; 755 '~Spare WB2[23].19'; 756 '~Spare WB2[23].20'; 757 '~Spare WB2[23].21'; 758 '~Spare WB2[23].22'; 759 '~Spare WB2[23].23'; 760 '~Spare WB2[23].24'; 761 '~Spare WB2[23].25'; 762 '~Spare WB2[23].26'; 763 '~Spare WB2[23].27'; 764 '~Spare WB2[23].28'; 765 '~Spare WB2[23].29'; 766 '~Spare WB2[23].30'; 767 '~Spare WB2[23].31'; 768 '~Spare WB2[24].0'; 769 '~Spare WB2[24].1'; 770 '~Spare WB2[24].2'; 771 '~Spare WB2[24].3'; 772 '~Spare WB2[24].4'; 773 '~Spare WB2[24].5'; 774 '~Spare WB2[24].6'; 775 '~Spare WB2[24].7'; 776 '~Spare WB2[24].8'; 777 '~Spare WB2[24].9'; 778 '~Spare WB2[24].10'; 779 '~Spare WB2[24].11'; 780 '~Spare WB2[24].12'; 781 '~Spare WB2[24].13'; 782 '~Spare WB2[24].14'; 783 '~Spare WB2[24].15'; 784 '~Spare WB2[24].16'; 785 '~Spare WB2[24].17'; 786 '~Spare WB2[24].18'; 787 '~Spare WB2[24].19'; 788 '~Spare WB2[24].20'; 789 '~Spare WB2[24].21'; 790 '~Spare WB2[24].22'; 791 '~Spare WB2[24].23'; 792 '~Spare WB2[24].24'; 793 '~Spare WB2[24].25'; 794 '~Spare WB2[24].26'; 795 '~Spare WB2[24].27'; 796 '~Spare WB2[24].28'; 797 '~Spare WB2[24].29'; 798 '~Spare WB2[24].30'; 799 '~Spare WB2[24].31'; 800 '~Spare WB2[25].0'; 801 '~Spare WB2[25].1'; 802 '~Spare WB2[25].2'; 803 '~Spare WB2[25].3'; 804 '~Spare WB2[25].4'; 805 '~Spare WB2[25].5'; 806 '~Spare WB2[25].6'; 807 '~Spare WB2[25].7'; 808 '~Spare WB2[25].8'; 809 '~Spare WB2[25].9'; 810 '~Spare WB2[25].10'; 811 '~Spare WB2[25].11'; 812 '~Spare WB2[25].12'; 813 '~Spare WB2[25].13'; 814 '~Spare WB2[25].14'; 815 '~Spare WB2[25].15'; 816 '~Spare WB2[25].16'; 817 '~Spare WB2[25].17'; 818 '~Spare WB2[25].18'; 819 '~Spare WB2[25].19'; 820 '~Spare WB2[25].20'; 821 '~Spare WB2[25].21'; 822 '~Spare WB2[25].22'; 823 '~Spare WB2[25].23'; 824 '~Spare WB2[25].24'; 825 '~Spare WB2[25].25'; 826 '~Spare WB2[25].26'; 827 '~Spare WB2[25].27'; 828 '~Spare WB2[25].28'; 829 '~Spare WB2[25].29'; 830 '~Spare WB2[25].30'; 831 '~Spare WB2[25].31'; 832 '~S001R11 Waiting Zone #1 Not Clear WB2[26].0'; 833 '~S001R11 Waiting Zone #2 Not Clear WB2[26].1'; 834 '~S001R11 Waiting Zone #3 Not Clear WB2[26].2'; 835 '~S001R11 Waiting Zone #4 Not Clear WB2[26].3'; 836 '~S001R11 Waiting Zone #5 Not Clear WB2[26].4'; 837 '~S001R11 Waiting Zone #6 Not Clear WB2[26].5'; 838 '~S001R11 Waiting Zone #7 Not Clear WB2[26].6'; 839 '~S001R11 Waiting Zone #8 Not Clear WB2[26].7'; 840 '~S001R11 Waiting Zone #9 Not Clear WB2[26].8'; 841 '~S001R11 Waiting Zone #10 Not Clear WB2[26].9'; 842 '~S001R11 Waiting Zone #11 Not Clear WB2[26].10'; 843 '~S001R11 Waiting Zone #12 Not Clear WB2[26].11'; 844 '~S001R11 Waiting Zone #13 Not Clear WB2[26].12'; 845 '~S001R11 Waiting Zone #14 Not Clear WB2[26].13'; 846 '~S001R11 Waiting Tip Dress Zone #1 Not Clear WB2[26].14'; 847 '~S001R11 Waiting Tip Dress Zone #2 Not Clear WB2[26].15'; 848 '~S001R11 Adjacent Robot xx-xx In Teach WB2[26].16'; 849 '~S001R11 Adjacent Robot xx-xx In Teach WB2[26].17'; 850 '~S001R11 Adjacent Robot xx-xx In Teach WB2[26].18'; 851 '~S001R11 Adjacent Robot xx-xx In Teach WB2[26].19'; 852 '~S001R11 Adjacent Robot xx-xx In Teach WB2[26].20'; 853 '~S001R11 Adjacent Robot xx-xx In Teach WB2[26].21'; 854 '~S001R11 Adjacent Robot xx-xx In Teach WB2[26].22'; 855 '~S001R11 Adjacent Robot xx-xx In Teach WB2[26].23'; 856 '~S001R11 Adjacent Robot xx-xx In Teach WB2[26].24'; 857 '~S001R11 Adjacent Robot xx-xx In Teach WB2[26].25'; 858 '~Spare WB2[26].26'; 859 '~Spare WB2[26].27'; 860 '~Spare WB2[26].28'; 861 '~S001R11 Robot Not Clear Of Fixture WB2[26].29'; 862 '~Spare WB2[26].30'; 863 '~Spare WB2[26].31'; 864 '~Spare WB2[27].0'; 865 '~Spare WB2[27].1'; 866 '~Spare WB2[27].2'; 867 '~Spare WB2[27].3'; 868 '~Spare WB2[27].4'; 869 '~Spare WB2[27].5'; 870 '~Spare WB2[27].6'; 871 '~Spare WB2[27].7'; 872 '~Spare WB2[27].8'; 873 '~Spare WB2[27].9'; 874 '~Spare WB2[27].10'; 875 '~Spare WB2[27].11'; 876 '~Spare WB2[27].12'; 877 '~Spare WB2[27].13'; 878 '~Spare WB2[27].14'; 879 '~Spare WB2[27].15'; 880 '~Spare WB2[27].16'; 881 '~Spare WB2[27].17'; 882 '~Spare WB2[27].18'; 883 '~Spare WB2[27].19'; 884 '~Spare WB2[27].20'; 885 '~Spare WB2[27].21'; 886 '~Spare WB2[27].22'; 887 '~Spare WB2[27].23'; 888 '~Spare WB2[27].24'; 889 '~Spare WB2[27].25'; 890 '~Spare WB2[27].26'; 891 '~Spare WB2[27].27'; 892 '~Spare WB2[27].28'; 893 '~Spare WB2[27].29'; 894 '~Spare WB2[27].30'; 895 '~Spare WB2[27].31'; 896 '~S001R11 Cycle Overtime WB2[28].0'; 897 '~S001R11 In Bypass WB2[28].1'; 898 '~S001R11 Battery Low WB2[28].2'; 899 '~S001R11 Servo Over Torque WB2[28].3'; 900 '~S001R11 Process Retry In Progress WB2[28].4'; 901 '~Spare WB2[28].5'; 902 '~S001R11 Robot Edit Occurred Ext App WB2[28].6'; 903 '~S001R11 Robot Input Simmed WB2[28].7'; 904 '~S001R11 Robot Output Simmed WB2[28].8'; 905 '~Spare WB2[28].9'; 906 '~Spare WB2[28].10'; 907 '~Spare WB2[28].11'; 908 '~Spare WB2[28].12'; 909 '~Spare WB2[28].13'; 910 '~Spare WB2[28].14'; 911 '~Spare WB2[28].15'; 912 '~S001R11F1B1.M.ModuleFlt - Externa App 1 I/O Module Warning WB2[28].16'; 913 '~S001R11F2B1.M.ModuleFlt - Externa App 2 I/O Module Warning WB2[28].17'; 914 '~S001R11F3B1.M.ModuleFlt - Externa App 3 I/O Module Warning WB2[28].18'; 915 '~Spare WB2[28].19'; 916 '~Spare WB2[28].20'; 917 '~Spare WB2[28].21'; 918 '~Spare WB2[28].22'; 919 '~Spare WB2[28].23'; 920 '~S001R11ES1 - S001R11 EtherNet Switch Port At Half Duplex WB2[28].24'; 921 '~S001R11ES1 - S001R11 EtherNet Switch Config Changes Not Saved WB2[28].25'; 922 '~S001R11ES1 - S001R11 EtherNet Switch Configuration Changed WB2[28].26'; 923 '~S001R11ES1 - S001R11 EtherNet Switch Port With Excessive Errors WB2[28].27'; 924 '~S001R11ES1 - S001R11 EtherNet Switch Port With Utilization Warning WB2[28].28'; 925 '~S001R11ES1 - S001R11 EtherNet Switch Changes Require Reboot WB2[28].29'; 926 '~Spare WB2[28].30'; 927 '~Spare WB2[28].31'; 928 '~Spare WB2[29].0'; 929 '~Spare WB2[29].1'; 930 '~S001R11 Servo Gun Tip Calib Request 1 WB2[29].2'; 931 '~S001R11 I-Available Warning 1 WB2[29].3'; 932 '~S001R11 Tip Dress Motor 1 Fault Bypassed WB2[29].4'; 933 '~S001R11 Tip Change Notice 1 WB2[29].5'; 934 '~S001R11 Bypass Tip Dresser 1 Selected WB2[29].6'; 935 '~S001R11 Auto Tip Changer Low 1 WB2[29].7'; 936 '~S001R11 Auto Tip Changer Empty 1 WB2[29].8'; 937 '~S001R11 Tip Wear Ratio Warning 1 - Touch Up Tip Dress Program WB2[29].9'; 938 '~S001R11 Stud Weld 1 Maintenance Reqd WB2[29].10'; 939 '~S001R11 Stud Weld 1 Low Stud Warning WB2[29].11'; 940 '~Spare WB2[29].12'; 941 '~S001R11 Rivet 1 Low Rivet Warning WB2[29].13'; 942 '~S001R11 Rivet 1 - Skip Once Initiated from Robot TP WB2[29].14'; 943 '~S001R11 Rivet 1 - Skip Remaining Initiated from Robot TP WB2[29].15'; 944 '~S001R11 Rivet 1 Preventive Maintenace Required WB2[29].16'; 945 '~S001R11 Rivet 1 Magazine Low WB2[29].17'; 946 '~S001R11 Tip Change 1 Bypassed WB2[29].18'; 947 '~S001R11 Mig Weld Fluid Level Low WB2[29].19'; 948 '~S001R11 Weld Ctrlr 1 Adaptive Mode Is Disabled WB2[29].20'; 949 '~S001R11 Tip Cutter 1 Warning WB2[29].21'; 950 '~S001R11 Rivet 1 Tape-Cut Required WB2[29].22'; 951 '~S001R11 Wire Feeder Motor Over Current WB2[29].23'; 952 '~Spare WB2[29].24'; 953 '~S001R11 Sealer Ctrlr 1 Minor Fault WB2[29].25'; 954 '~S001R11 Sealer Ctrlr 1 Required Rezeroing WB2[29].26'; 955 '~S001R11 Loaded To Average WB2[29].27'; 956 '~S001R11 Vision Process Aborted WB2[29].28'; 957 '~S001R11 Vision System Trending WB2[29].29'; 958 '~S001R11 Vision Out Of Tolerance WB2[29].30'; 959 '~Spare WB2[29].31'; 960 '~Spare WB2[30].0'; 961 '~Spare WB2[30].1'; 962 '~S001R11 Servo Gun Tip Calib Request 2 WB2[30].2'; 963 '~S001R11 I-Available Warning 2 WB2[30].3'; 964 '~S001R11 Tip Dress Motor 2 Fault Bypassed WB2[30].4'; 965 '~S001R11 Tip Change Notice 2 WB2[30].5'; 966 '~S001R11 Bypass Tip Dresser 2 Selected WB2[30].6'; 967 '~S001R11 Auto Tip Changer Low 2 WB2[30].7'; 968 '~S001R11 Auto Tip Changer Empty 2 WB2[30].8'; 969 '~S001R11 Tip Wear Ratio Warning 2 - Touch Up Tip Dress Program WB2[30].9'; 970 '~S001R11 Stud Weld 2 Maintenance Reqd WB2[30].10'; 971 '~S001R11 Stud Weld 2 Low Stud Warning WB2[30].11'; 972 '~Spare WB2[30].12'; 973 '~S001R11 Rivet 2 Low Rivet Warning WB2[30].13'; 974 '~S001R11 Rivet 2 - Skip Once Initiated from Robot TP WB2[30].14'; 975 '~S001R11 Rivet 2 - Skip Remaining Initiated from Robot TP WB2[30].15'; 976 '~S001R11 Rivet 2 Preventive Maintenace Required WB2[30].16'; 977 '~S001R11 Rivet 2 Magazine Low WB2[30].17'; 978 '~S001R11 Tip Change 2 Bypassed WB2[30].18'; 979 '~S001R11 Laser Dirty Glass Warning WB2[30].19'; 980 '~S001R11 Weld Ctrlr 2 Adaptive Mode Is Disabled WB2[30].20'; 981 '~S001R11 Tip Cutter 2 Warning WB2[30].21'; 982 '~S001R11 Rivet 2 Tape-Cut Required WB2[30].22'; 983 '~S001R11 Mig Tip Nozzel Replacement Warning WB2[30].23'; 984 '~S001R11 Mig Tip Nozzel Replacement Required WB2[30].24'; 985 '~S001R11 Sealer Ctrlr 2 Minor Fault WB2[30].25';